
                   //PathData - command - valueFlags
                   //====================================================================================================================================
                   // also copy flagMode to pathDataPreBuf for use in specific case of waitFlag
                   FOR #tempFlagCtr := 1 TO "LKINCTRL_NO_OF_CMD_VALUEFLAGS" DO
                       #pathDataPreBuf.commands[#pathDataPreBuf.addPointer].valueFlags[#tempFlagCtr] := #statPathDataCommand.valueFlags[#tempFlagCtr];
                       // // change flagMode 3 to flagMode 2 as functionality is equal
                       // check for cmd to be flagOnly cmd
                       // check for cmd to implement flag and flagMode to be flagMode 3
                       IF #pathDataPreBuf.commands[#pathDataPreBuf.addPointer].cmdType = "LKINCTRL_CMD_FLAG_ONLY"
                           AND #pathDataPreBuf.commands[#pathDataPreBuf.addPointer].valueFlags[#tempFlagCtr].flag <> -1
                           AND #pathDataPreBuf.commands[#pathDataPreBuf.addPointer].valueFlags[#tempFlagCtr].flagMode = 3
                       THEN
                           // change flagMode 3 to flagMode 2
                           #pathDataPreBuf.commands[#pathDataPreBuf.addPointer].valueFlags[#tempFlagCtr].flagMode := 2;
                       END_IF;
                   END_FOR;

                   // skip lastPos calculation in case of wait time execution ==> old lastPos will be correct ==> use separation of config / motion cmd (flagOnly)
                   IF #statCmdIsMotionCmd THEN
                       //------------------------------------------------------------------------------------------
                       // Transform statLastPos into correct CS
                       //------------------------------------------------------------------------------------------
                       // TODO: Integrate InverseKinTrans into FC LKinCtrl_FrameTrans ?
                       IF #statPathDataCommand.cmdCoordinates.coordSystem = "CS_MCS"
                           AND #statCoordSystemOld <> "CS_MCS"
                       THEN
                           // Transform lastPos to MCS 
                           #instMC_InverseKinematicsTransformation(AxesGroup := #to_Kinematics,
                                                                   Enable := TRUE,
                                                                   Position := #statLastPos,
                                                                   CoordSystem := #statCoordSystemOld,
                                                                   LinkConstellation := #statLinkConstellation,
                                                                   ErrorId => #tempRetVal,
                                                                   AxesPosition => #statLastPos);

                       ELSIF #statPathDataCommand.cmdCoordinates.coordSystem <> "CS_MCS"
                           AND #statCoordSystemOld = "CS_MCS"
                       THEN
                           // Transform lastPos to target CS
                           #instMC_KinematicsTransformation(AxesGroup := #to_Kinematics,
                                                            Enable := TRUE,
                                                            AxesPosition := #statLastPos,
                                                            CoordSystem := #statPathDataCommand.cmdCoordinates.coordSystem,
                                                            ErrorId => #tempRetVal,
                                                            Position => #statLastPos,
                                                            LinkConstellation => #statLinkConstellation);

                       ELSE
                           // FR 26.03.2020: Updated FrameTrans 
                           // Transform LastPos to correct CS
                           "LKinCtrl_FrameTrans"(coordSystem := #statPathDataCommand.cmdCoordinates.coordSystem, // Actual/Target CS
                                                 coordSystemOld := #statCoordSystemOld, // Last CS
                                                 OCSFrames := #OCSFrames, // OCS frames
                                                 position := #statLastPos); // Position to be transformed
                       END_IF;

                       // Check if KinTrans FBs returned no error
                       IF #tempRetVal = 16#0 THEN
                           // Update old CS
                           #statCoordSystemOld := #statPathDataCommand.cmdCoordinates.coordSystem;

                           //------------------------------------------------------------------------------------------
                           // Update linkConstellation
                           //------------------------------------------------------------------------------------------
                           // LinkConstellation can only be set at sPTP command in WCS/OCS
                           IF #statPathDataCommand.cmdCoordinates.coordSystem <> "CS_MCS"
                               AND #statPathDataCommand.cmdParameters.moveDirectParameters.linkConstellation <> 16#FFFF_FFFF
                               AND (#statPathDataCommand.cmdType = "LKINCTRL_MC_MOVEDIRECTABS"
                               OR #statPathDataCommand.cmdType = "LKINCTRL_MC_MOVEDIRECTREL")
                           THEN
                               // LinkConstellation is changed
                               #statLinkConstellation := DWORD_TO_DINT(#statPathDataCommand.cmdParameters.moveDirectParameters.linkConstellation);
                           END_IF;

                           //------------------------------------------------------------------------------------------
                           // Update PositionMode
                           //------------------------------------------------------------------------------------------
                           // PositionMode is only valid for absolute SPTP command in WCS/OCS
                           IF #statPathDataCommand.cmdCoordinates.coordSystem <> "CS_MCS"
                               AND #statPathDataCommand.cmdParameters.moveDirectParameters.positionMode = 2 // Relative A coordinate
                               AND #statPathDataCommand.cmdType = "LKINCTRL_MC_MOVEDIRECTABS"
                           THEN
                               // Calc correct orientation position
                               #statLastPos[4] := #statLastPos[4] + #statPathDataCommand.cmdCoordinates.cartesianPosition.a;
                           END_IF;

                           //------------------------------------------------------------------------------------------
                           // ParameterValid bit check
                           //------------------------------------------------------------------------------------------
                           // added FR: 2020/04/03
                           "LKinCtrl_EvaluateParamValidBits"(parameterValidBits := #statParameterValid,
                                                             lastPos := #statLastPos,
                                                             errorMessage => #statDebugMessage,
                                                             command := #statPathDataCommand);

                           // Caclulation of resulting last position after command
                           //====================================================================================================================================
                           #statRetValLastPos := "LKinCtrl_CalcResultingPos"(cmdType := #statPathDataCommand.cmdType,
                                                                             cartesianPos := #statPathDataCommand.cmdCoordinates.cartesianPosition,
                                                                             circleParameters := #statPathDataCommand.cmdParameters.circleParameters,
                                                                             errorMessage => #statDebugMessage,
                                                                             lastPos := #statLastPos,
                                                                             lastAuxPoint := #statAuxPoint);

                           // check for error in last position calculation
                           IF #statRetValLastPos <> 16#0 THEN
                               // set error status
                               #statErrorAutoCleared := TRUE;
                               #statStatus := #ERR_LASTPOS_CALCULATION;
                           END_IF;

                       ELSE
                           // Error in KinTrans FBs
                           // set error status
                           #statErrorAutoCleared := TRUE;
                           #statStatus := #tempRetVal;
                       END_IF;

                   END_IF;

                   // PathData Blending at start of path
                   IF (#statPathDataPointers.retrievePointer = 1) AND
                       (#initPathTransition = 1)
                   THEN
                       #pathDataPreBuf.commands[#pathDataPreBuf.addPointer].cmdParameters.bufferMode := #initBufferMode;
                       #pathDataPreBuf.commands[#pathDataPreBuf.addPointer].cmdParameters.transitionParameters := #initTransitionParameter;
                   END_IF;

                   // increment PathDataPreBuf addPointer for next copy procedure
                   // also implement restart of pointer (1..constant)
                   IF #pathDataPreBuf.addPointer < "LKINCTRL_NO_OF_PATHDATA_PREBUFFER_ELEMENTS" THEN
                       #pathDataPreBuf.addPointer += 1;
                   ELSE
                       #pathDataPreBuf.addPointer := 1;
                       #pathDataPreBuf.addPointerRestarted := TRUE;
                   END_IF;
               END_REGION COPY_CMD_REGULAR

               // Go to copy cmd
               #statStateMachine := #GET_CMD;
           END_IF;


           // =======================================================================================================  
           // Contour offset is handled in the following regions / states
           // =======================================================================================================  
           REGION CONTOUR_OFFSET

               // STATE: CHECK_NEXT_CMD
               // =======================================================================================================  
               // CHECK_NEXT_CMD: Check next command for contour offset (#statPathCmdOffCompIn.nextCommand)
               // Next state: OFFSET_CALC / SEARCH_NBO
               IF #statStateMachine = #CHECK_NEXT_CMD THEN
                   REGION CHECK_NEXT_CMD
                       // Check if current command has length 0.0 --> Copy without contour offset
                       // else use as nextCmd & search NBO
                       // Transform lastPos to correct CS
                       "LKinCtrl_FrameTrans"(coordSystem := #statPathDataCommand.cmdCoordinates.coordSystem,
                                             coordSystemOld := #statCoordSystemOld,
                                             OCSFrames := #OCSFrames,
                                             position := #statLastPos);

                       // Update old CS
                       #statCoordSystemOld := #statPathDataCommand.cmdCoordinates.coordSystem;

                       // ParameterValid bit check
                       "LKinCtrl_EvaluateParamValidBits"(parameterValidBits := #statParameterValid,
                                                         lastPos := #statLastPos,
                                                         errorMessage => #statDebugMessage,
                                                         command := #statPathDataCommand);

                       // implement CM3 ==> CM1 conversion here
                       #statRetValCircModeConv := "LKinCtrl_ConvCircMode3To1"(coordinates := #statPathDataCommand.cmdCoordinates.cartesianPosition,
                                                                              errorMessage => #statDebugMessage,
                                                                              lastPos := #statLastPos,
                                                                              cmdType := #statPathDataCommand.cmdType,
                                                                              circleParameters := #statPathDataCommand.cmdParameters.circleParameters);

                       // Check if cmd has 0.0 length
                       "LKinCtrl_CheckForCmdLengthZero"(lastPos := #statLastPos,
                                                        commandLengthIsZero => #tempCmdLengthIsZero,
                                                        command := #statPathDataCommand);

                       // check for command length to be zero
                       IF #tempCmdLengthIsZero = FALSE THEN
                           // Comd is not length 0.0

                           // Calc resulting pos to use for searching NBO
                           #statRetValLastPos := "LKinCtrl_CalcResultingPos"(cmdType := #statPathDataCommand.cmdType,
                                                                             cartesianPos := #statPathDataCommand.cmdCoordinates.cartesianPosition,
                                                                             circleParameters := #statPathDataCommand.cmdParameters.circleParameters,
                                                                             errorMessage => #statDebugMessage,
                                                                             lastAuxPoint := #statAuxPoint,
                                                                             lastPos := #statLastPos);


                           // Use as next cmd
                           // set first condition bit to abort loop
                           #tempValidNextCmdFound := TRUE;
                           #statDebugNextCmdFound := #statPathDataPointers.retrievePointer;

                           // check for command to be END_OFFSET_COMP command
                           IF #statPathDataCommand.cmdType = "LKINCTRL_CONFIG_END_OFFSET_COMP"
                               OR #statPathDataCommand.cmdType = -1
                           THEN
                               // transfer no command for end of compensation
                               #statPathCmdOffCompIn.nextCommand.cmdType := -1;
                               // transfer no command for end of compensation
                               #statPathCmdOffCompIn.nextButOneCommand.cmdType := -1;
                               #tempValidNextButOneCmdFound := TRUE;
                               // Go to next state --> No need to search NBO
                               #statStateMachine := #OFFSET_CALC;
                           ELSE
                               // copy 'next' cmd to next(ButOne)Command input
                               #statPathCmdOffCompIn.nextCommand := #statPathDataCommand;
                               // Go to next state
                               #statStateMachine := #SEARCH_NBO;
                           END_IF;

                       ELSE
                           // command has no length --> RelCmd with 0.0 or AbsCmd with same target
                           // copy command as usual without calling any contour offset calculation functions
                           REGION COPY_LENGTH_0_CMD
                               //PathData - command - cmdType
                               #pathDataPreBuf.commands[#pathDataPreBuf.addPointer].cmdType := #statPathDataCommand.cmdType;

                               //PathData - command - cmdID
                               #pathDataPreBuf.commands[#pathDataPreBuf.addPointer].cmdID := #statPathDataPointers.retrievePointer + #statNoRestarts * INT_TO_DINT("LKINCTRL_NO_OF_PATHDATA_ELEMENTS_ADVANCED");

                               //PathData - command - cmdName
                               #pathDataPreBuf.commands[#pathDataPreBuf.addPointer].cmdName := #statPathDataCommand.cmdName;

                               //PathData - command - cmdCoordinates
                               //====================================================================================================================================
                               //PathData - command - cmdCoordinates - absolutePosition[1..4]
                               IF #statOffsetCompFirstCmd = FALSE AND #statPathDataCommand.cmdType = "LKINCTRL_MC_MOVELINEARABS" THEN
                                   // Use compensated coordinates for multiple zero length commands in a row
                                   #pathDataPreBuf.commands[#pathDataPreBuf.addPointer].cmdCoordinates.absolutePosition[1] := #statPathCmdOffCompIn.currentPos.positionAbsoluteRadComp.x;
                                   #pathDataPreBuf.commands[#pathDataPreBuf.addPointer].cmdCoordinates.absolutePosition[2] := #statPathCmdOffCompIn.currentPos.positionAbsoluteRadComp.y;
                                   #pathDataPreBuf.commands[#pathDataPreBuf.addPointer].cmdCoordinates.absolutePosition[3] := #statPathCmdOffCompIn.currentPos.positionAbsoluteRadComp.z;
                                   #pathDataPreBuf.commands[#pathDataPreBuf.addPointer].cmdCoordinates.absolutePosition[4] := #statPathCmdOffCompIn.currentPos.positionAbsoluteRadComp.a;
                               ELSE
                                   #pathDataPreBuf.commands[#pathDataPreBuf.addPointer].cmdCoordinates.absolutePosition[1] := #statPathDataCommand.cmdCoordinates.cartesianPosition.x;
                                   #pathDataPreBuf.commands[#pathDataPreBuf.addPointer].cmdCoordinates.absolutePosition[2] := #statPathDataCommand.cmdCoordinates.cartesianPosition.y;
                                   #pathDataPreBuf.commands[#pathDataPreBuf.addPointer].cmdCoordinates.absolutePosition[3] := #statPathDataCommand.cmdCoordinates.cartesianPosition.z;
                                   #pathDataPreBuf.commands[#pathDataPreBuf.addPointer].cmdCoordinates.absolutePosition[4] := #statPathDataCommand.cmdCoordinates.cartesianPosition.a;
                               END_IF;

                               //PathData - command - cmdCoordinates - coordSystem
                               #pathDataPreBuf.commands[#pathDataPreBuf.addPointer].cmdCoordinates.coordSystem := #statPathDataCommand.cmdCoordinates.coordSystem;

                               //PathData - command - cmdParameters
                               //====================================================================================================================================
                               //PathData - command - cmdParameters - pathDynamics
                               #pathDataPreBuf.commands[#pathDataPreBuf.addPointer].cmdParameters.pathDynamics := #statPathDataCommand.cmdParameters.pathDynamics;

                               //PathData - command - cmdParameters - orientationDirection
                               #pathDataPreBuf.commands[#pathDataPreBuf.addPointer].cmdParameters.orientationDirection := #statPathDataCommand.cmdParameters.orientationDirection;

                               //PathData - command - cmdParameters - bufferMode
                               #pathDataPreBuf.commands[#pathDataPreBuf.addPointer].cmdParameters.bufferMode := #statPathDataCommand.cmdParameters.bufferMode;

                               //PathData - command - cmdParameters - transitionParameters
                               #pathDataPreBuf.commands[#pathDataPreBuf.addPointer].cmdParameters.transitionParameters[1] := #statPathDataCommand.cmdParameters.transitionParameters[1];

                               //PathData - command - cmdParameters - dynamicAdaption
                               #pathDataPreBuf.commands[#pathDataPreBuf.addPointer].cmdParameters.dynamicAdaption := #statPathDataCommand.cmdParameters.dynamicAdaption;

                               //PathData - command - setFlags
                               //====================================================================================================================================
                               // also copy flagMode to pathDataPreBuf for use in specific case of waitFlag
                               FOR #tempFlagCtr := 1 TO "LKINCTRL_NO_OF_CMD_SETFLAGS" DO
                                   #pathDataPreBuf.commands[#pathDataPreBuf.addPointer].setFlags[#tempFlagCtr] := #statPathDataCommand.setFlags[#tempFlagCtr];
                                   // // change flagMode 3 to flagMode 2 as functionality is equal
                                   // check for cmd to be flagOnly cmd
                                   // check for cmd to implement flag and flagMode to be flagMode 3
                                   IF #pathDataPreBuf.commands[#pathDataPreBuf.addPointer].cmdType = "LKINCTRL_CMD_FLAG_ONLY"
                                       AND #pathDataPreBuf.commands[#pathDataPreBuf.addPointer].setFlags[#tempFlagCtr].flag <> -1
                                       AND #pathDataPreBuf.commands[#pathDataPreBuf.addPointer].setFlags[#tempFlagCtr].flagMode = 3
                                   THEN
                                       // change flagMode to flagMode 1
                                       #pathDataPreBuf.commands[#pathDataPreBuf.addPointer].setFlags[#tempFlagCtr].flagMode := 2;
                                   END_IF;
                               END_FOR;

                               //PathData - command - valueFlags
                               //====================================================================================================================================
                               // also copy flagMode to pathDataPreBuf for use in specific case of waitFlag
                               FOR #tempFlagCtr := 1 TO "LKINCTRL_NO_OF_CMD_VALUEFLAGS" DO
                                   #pathDataPreBuf.commands[#pathDataPreBuf.addPointer].valueFlags[#tempFlagCtr] := #statPathDataCommand.valueFlags[#tempFlagCtr];
                                   // // change flagMode 3 to flagMode 2 as functionality is equal
                                   // check for cmd to be flagOnly cmd
                                   // check for cmd to implement flag and flagMode to be flagMode 3
                                   IF #pathDataPreBuf.commands[#pathDataPreBuf.addPointer].cmdType = "LKINCTRL_CMD_FLAG_ONLY"
                                       AND #pathDataPreBuf.commands[#pathDataPreBuf.addPointer].valueFlags[#tempFlagCtr].flag <> -1
                                       AND #pathDataPreBuf.commands[#pathDataPreBuf.addPointer].valueFlags[#tempFlagCtr].flagMode = 3
                                   THEN
                                       // change flagMode to flagMode 1
                                       #pathDataPreBuf.commands[#pathDataPreBuf.addPointer].valueFlags[#tempFlagCtr].flagMode := 2;
                                   END_IF;

                               END_FOR;

                               // increase addPointer after copy of command for next command
                               IF #pathDataPreBuf.addPointer < "LKINCTRL_NO_OF_PATHDATA_PREBUFFER_ELEMENTS" THEN
                                   #pathDataPreBuf.addPointer += 1;
                               ELSE
                                   #pathDataPreBuf.addPointer := 1;
                                   #pathDataPreBuf.addPointerRestarted := TRUE;
                               END_IF;

                           END_REGION COPY_REL_0_CMD

                           // Go to next state
                           #statStateMachine := #OFFSET_CALC;

                       END_IF;
                   END_REGION CHECK_NEXT_CMD
               END_IF;


               // STATE: SEARCH_NBO
               // =======================================================================================================  
               // SEARCH_NBO: Search forward in path data for contour offset next but one command (#statPathCmdOffCompIn.nextButOneCommand)
               // Next state: OFFSET_CALC
               IF #statStateMachine = #SEARCH_NBO THEN
                   REGION SEARCH_NBO
                       // find valid nextCmd and nextButOneCmd (input) data
                       // ---------------------------------------------------
                       // Init last pos and old coord system
                       #statNBOLastPos := #statLastPos;
                       #tempNBOCoordSystemOld := #statCoordSystemOld;

                       IF #statSearchNBOAborted = FALSE THEN
                           // initially set pointer increase counter to 1
                           #statRetrievePointerIncCtr := 1;
                       ELSE
                           // Reset abort bit but keep RetreivePointerIncCounter the same
                           #statSearchNBOAborted := FALSE;
                       END_IF;

                       // Use repeat to search in path data for next valid command
                       REPEAT

                           // Check pointers also for not ringBuffer or ignore add pointer
                           // Added FR 22.05.2019
                           IF #statPathDataPointers.ignoreAddPointer THEN
                               // No ring buffer
                               // Check index to be lower than max path data length 
                               IF #statPathDataType = "LKINCTRL_PATHDATA_TYPE_REDUCED" THEN
                                   #tempIndexOk := #statPathDataPointers.retrievePointer + #statRetrievePointerIncCtr <= "LKINCTRL_NO_OF_PATHDATA_ELEMENTS_REDUCED";
                               ELSIF #statPathDataType = "LKINCTRL_PATHDATA_TYPE_NORMAL" THEN
                                   #tempIndexOk := #statPathDataPointers.retrievePointer + #statRetrievePointerIncCtr <= "LKINCTRL_NO_OF_PATHDATA_ELEMENTS";
                               ELSIF #statPathDataType = "LKINCTRL_PATHDATA_TYPE_ADVANCED" THEN
                                   #tempIndexOk := #statPathDataPointers.retrievePointer + #statRetrievePointerIncCtr <= "LKINCTRL_NO_OF_PATHDATA_ELEMENTS_ADVANCED";
                               END_IF;
                           ELSE
                               // Ring buffer
                               // Added JR 13.05.2019 
                               // If index overflows then calc offset to point to first index
                               IF #statPathDataPointers.retrievePointer + #statRetrievePointerIncCtr > "LKINCTRL_NO_OF_PATHDATA_ELEMENTS_ADVANCED" THEN
                                   // Set statRetrievePointerIncCtr
                                   #statRetrievePointerIncCtr := 1 - #statPathDataPointers.retrievePointer;
                               END_IF;

                               // Condition if (#statPathDataPointers.retrievePointer + #statRetrievePointerIncCtr) > 1
                               #tempIndexOk :=
                               ((#statPathDataPointers.retrievePointer + #statRetrievePointerIncCtr) <= #statPathDataPointers.addPointer)
                               OR (((#statPathDataPointers.retrievePointer + #statRetrievePointerIncCtr) > #statPathDataPointers.addPointer)
                               AND #statPathDataPointers.addPointerRestarted);
                           END_IF;

                           // Copy path data command
                           // 2019.03.28 FR: Get last command
                           IF (#statPathDataPointers.retrievePointer + #statRetrievePointerIncCtr) >= 1
                               AND #tempIndexOk
                           THEN
                               // Get path data command and previous path data command
                               #tempRetVal := "LKinCtrl_GetPathDataCmd"(pathDataType := #statPathDataType,
                                                                        index := #statPathDataPointers.retrievePointer + #statRetrievePointerIncCtr,
                                                                        pathDataReduced := #tempPathData_reduced,
                                                                        pathData := #tempPathData,
                                                                        pathDataAdvanced := #tempPathData_advanced,
                                                                        pathDataCommand => #statPathCmdNBOCheck,
                                                                        parameterValid => #tempParameterValidNBO);


                               // Check if index is not ok and not ring buffer
                               // --> End of path data is reached and Next or NBO was not found 
                               // --> Set the corresponding cmd to -1 to end offset correctly 
                           ELSIF #tempIndexOk = FALSE
                               AND #statPathDataPointers.ignoreAddPointer
                           THEN
                               IF #tempValidNextCmdFound THEN
                                   // set NBO to -1
                                   // transfer no command for end of compensation
                                   #statPathCmdOffCompIn.nextButOneCommand.cmdType := -1;
                                   #tempValidNextButOneCmdFound := TRUE;
                               ELSE
                                   // set Next and NBO to -1
                                   // transfer no command for end of compensation
                                   #statPathCmdOffCompIn.nextCommand.cmdType := -1;
                                   #tempValidNextCmdFound := TRUE;
                                   // transfer no command for end of compensation
                                   #statPathCmdOffCompIn.nextButOneCommand.cmdType := -1;
                                   #tempValidNextButOneCmdFound := TRUE;
                               END_IF;
                               // Exit repeat
                               EXIT;

                               // Index is not valid and ringbuffer active --> Check for new command 
                           ELSE
                               // Exit repeat loop and check again in next cycle
                               // memorize abort
                               #statSearchNBOAborted := TRUE;
                               EXIT;
                           END_IF;

                           // preCheck sequence for comamnd to have length of zero
                           #tempCmdLengthIsZero := FALSE;

                           // Command was copied --> Check if valid for NBO
                           IF #statPathCmdNBOCheck.cmdActivated THEN
                               // Valid
                               // Check for length 0.0
                               // Transform lastPos to correct CS
                               "LKinCtrl_FrameTrans"(coordSystem := #statPathCmdNBOCheck.cmdCoordinates.coordSystem,
                                                     coordSystemOld := #tempNBOCoordSystemOld,
                                                     OCSFrames := #OCSFrames,
                                                     position := #statNBOLastPos);

                               // Update old CS
                               #tempNBOCoordSystemOld := #statPathCmdNBOCheck.cmdCoordinates.coordSystem;

                               // ParameterValid bit check
                               "LKinCtrl_EvaluateParamValidBits"(parameterValidBits := #tempParameterValidNBO,
                                                                 lastPos := #statNBOLastPos,
                                                                 errorMessage => #statDebugMessage,
                                                                 command := #statPathCmdNBOCheck);

                               // implement CM3 ==> CM1 conversion here
                               #statRetValCircModeConv := "LKinCtrl_ConvCircMode3To1"(coordinates := #statPathCmdNBOCheck.cmdCoordinates.cartesianPosition,
                                                                                      errorMessage => #statDebugMessage,
                                                                                      lastPos := #statNBOLastPos,
                                                                                      cmdType := #statPathCmdNBOCheck.cmdType,
                                                                                      circleParameters := #statPathCmdNBOCheck.cmdParameters.circleParameters);

                               // Check if cmd has 0.0 length
                               "LKinCtrl_CheckForCmdLengthZero"(lastPos := #statNBOLastPos,
                                                                commandLengthIsZero => #tempCmdLengthIsZero,
                                                                command := #statPathCmdNBOCheck);

                               IF #tempCmdLengthIsZero = FALSE THEN
                                   // Has length
                                   // Check if valid
                                   // set condition bit to abort loop
                                   #tempValidNextButOneCmdFound := TRUE;
                                   #statDebugNextButOneCmdFound := #statPathDataPointers.retrievePointer + #statRetrievePointerIncCtr;

                                   // check for command to be END_OFFSET_COMP command
                                   IF #statPathCmdNBOCheck.cmdType = "LKINCTRL_CONFIG_END_OFFSET_COMP"
                                       OR #statPathCmdNBOCheck.cmdType = -1
                                   THEN
                                       // transfer no command for end of compensation
                                       #statPathCmdOffCompIn.nextButOneCommand.cmdType := -1;
                                   ELSE
                                       // copy 'next' cmd to nextButOneCommand input
                                       #statPathCmdOffCompIn.nextButOneCommand := #statPathCmdNBOCheck;
                                   END_IF;
                               ELSE
                                   // Is 0.0 length cmd --> Not valid for NBO --> Search continues
                                   // increase set pointer increase counter to check next element
                                   #statRetrievePointerIncCtr += 1;
                               END_IF;

                           ELSE
                               // Cmd deactivated --> Not valid
                               // increase set pointer increase counter to check next element
                               #statRetrievePointerIncCtr += 1;
                           END_IF;

                       UNTIL #tempValidNextButOneCmdFound END_REPEAT;

                       // If both cmds were found and no abort then go to offset calc
                       IF #tempValidNextButOneCmdFound AND NOT #statSearchNBOAborted THEN
                           // Go to OffsetCalc
                           #statStateMachine := #OFFSET_CALC;

                           // reset variable for first offset command
                           #statOffsetCompFirstCmd := FALSE;
                       END_IF;
                   END_REGION SEARCH_NBO
               END_IF;

               // STATE: OFFSET_CMD
               // =======================================================================================================   
               // OFFSET_CMD: Copy offset command
               IF #statStateMachine = #OFFSET_CALC THEN
                   REGION OFFSET_CALC
                       // Offset Compensation Calculation
                       //====================================================================================================================================
                       // prepare data for offset calculation ==> only use original commands (source Pathdata !)

                       // check for command length not to be zero
                       IF #tempCmdLengthIsZero = FALSE THEN

                           // run offset caclulation
                           #statRetValOffsetComp := "LKinCtrl_OffsetContour"(toolLength := #statToolLength,
                                                                             toolRadius := #statToolRadius,
                                                                             pathPlane := #statPathPlane,
                                                                             compensationDirection := #statCompDirection,
                                                                             pathDataIn := #statPathCmdOffCompIn,
                                                                             pathDataOut := #statPathCmdOffCompOut);

                           // check for errors in offset compensation calculation
                           IF #statRetValOffsetComp.returnValue <> 16#0 THEN
                               #statErrorAutoCleared := TRUE;
                               #statStatus := #statRetValOffsetComp.returnValue;
                           ELSE
                               // use nextPositionAbsolute from last calc as currentPositionAbsolute for next calc
                               #statPathCmdOffCompIn.currentPos.positionAbsolute := #statPathCmdOffCompOut.nextPositionAbsolute;
                               #statPathCmdOffCompIn.currentPos.positionAbsoluteRadComp := #statPathCmdOffCompOut.nextPositionAbsoluteRadComp;

                               // use results of offset compensation calculation
                               // check for compensated nextCmd to be available
                               IF #statPathCmdOffCompOut.nextCommand.cmdType <> -1 THEN
                                   //PathData - command - cmdID
                                   #pathDataPreBuf.commands[#pathDataPreBuf.addPointer].cmdID := #statPathDataPointers.retrievePointer + #statNoRestarts * INT_TO_DINT("LKINCTRL_NO_OF_PATHDATA_ELEMENTS_ADVANCED");

                                   // copy next cmd data (OUT) - compensated (new calculated data)
                                   "LKinCtrl_ConvElements_PathDataToPathData_PreBuf"(copyCompensatedParametes := TRUE,
                                                                                     copyTransitionParameters := FALSE, //true ,
                                                                                     copyFlags := TRUE,
                                                                                     pathDataElement := #statPathCmdOffCompOut.nextCommand,
                                                                                     pathDataPreBufElement := #pathDataPreBuf.commands[#pathDataPreBuf.addPointer],
                                                                                     pathDataName := #statPathDataName);

                                   // Added FR 22.05.2019: Set ParameterValid bits true
                                   FOR #tempCtr := 1 TO "LKINCTRL_NO_OF_VALID_BITS" DO
                                       #pathDataPreBuf.commands[#pathDataPreBuf.addPointer].parameterValid[#tempCtr] := TRUE;
                                   END_FOR;

                                   // increase addPointer after copy of command for next command
                                   IF #pathDataPreBuf.addPointer < "LKINCTRL_NO_OF_PATHDATA_PREBUFFER_ELEMENTS" THEN
                                       #pathDataPreBuf.addPointer += 1;
                                   ELSE
                                       #pathDataPreBuf.addPointer := 1;
                                       #pathDataPreBuf.addPointerRestarted := TRUE;
                                   END_IF;

                                   // write transitionParameters of nextButOneCmd result to next but one command
                                   #pathDataPreBuf.commands[#pathDataPreBuf.addPointer].cmdParameters.transitionParameters := #statPathCmdOffCompOut.nextButOneCommand.transitionParameter;
                               ELSE
                                   ; // Invalid command -> nothing to copy
                               END_IF;

                               // check if there is an additional intermediate command
                               IF (#statPathCmdOffCompOut.intermediateCommand.cmdType > 0) THEN

                                   // copy intermediate cmd to PathData_PreBuf - no flags
                                   "LKinCtrl_ConvElements_PathDataToPathData_PreBuf"(copyCompensatedParametes := TRUE,
                                                                                     copyTransitionParameters := FALSE,
                                                                                     copyFlags := FALSE,
                                                                                     pathDataElement := #statPathCmdOffCompOut.intermediateCommand,
                                                                                     pathDataPreBufElement := #pathDataPreBuf.commands[#pathDataPreBuf.addPointer],
                                                                                     pathDataName := #statPathDataName);

                                   //PathData - command - cmdID
                                   // set intermediate commands cmdID to cmdID of following command ==> flag handling similar to transitionParameter
                                   #pathDataPreBuf.commands[#pathDataPreBuf.addPointer].cmdID := (#statPathDataPointers.retrievePointer + 1) + #statNoRestarts * INT_TO_DINT("LKINCTRL_NO_OF_PATHDATA_ELEMENTS_ADVANCED");

                                   // added FR: 11.07.2019: Set ParameterValid bits true
                                   FOR #tempCtr := 1 TO "LKINCTRL_NO_OF_VALID_BITS" DO
                                       #pathDataPreBuf.commands[#pathDataPreBuf.addPointer].parameterValid[#tempCtr] := TRUE;
                                   END_FOR;

                                   // mark intermediate commands to except them from flag for remaining distance
                                   #pathDataPreBuf.commands[#pathDataPreBuf.addPointer].isIntermediateCmd := TRUE;

                                   // increase addPointer after copy of command for next command
                                   IF #pathDataPreBuf.addPointer < "LKINCTRL_NO_OF_PATHDATA_PREBUFFER_ELEMENTS" THEN
                                       #pathDataPreBuf.addPointer += 1;
                                   ELSE
                                       #pathDataPreBuf.addPointer := 1;
                                       #pathDataPreBuf.addPointerRestarted := TRUE;
                                   END_IF;

                               ELSE
                                   ; // No intermediate cmd -> do nothing
                               END_IF;
                           END_IF;

                       ELSE
                           ; // do nothing --> Command was already copied
                       END_IF;

                   END_REGION OFFSET_CALC

                   // Go to copy cmd
                   #statStateMachine := #GET_CMD;
               END_IF;
           END_REGION CONTOUR_OFFSET

       END_REGION PATHDATA_PREBUFFERING


       REGION PATHDATA_PREBUFFERED_COMPLETELY
           // STATE: PATHDATA_PREBUFFERED_COMPLETELY
           // =======================================================================================================      
           // PATHDATA_PREBUFFERED_COMPLETELY: Disabling, e.g. closing connections, etc.
           IF #statStateMachine = #PATHDATA_PREBUFFERED_COMPLETELY
               // AND #statDebugState = TRUE
           THEN

               // reset  variable for single step debugging of states
               #statDebugState := FALSE;

               // Added FR 2019.03.28 // Reworked 08.04.2020
               // REGION GET_LAST_CMD_TYPE
               //
               // Always get last cmd id from preBuffered
               // --> Deactivated commands do not appear in preBuffered anyway
               // --> No need to check config cmds as they also do not appear --> Output LastCmdIsConfigCmd is not even needed / used in MovePath
               // --> Last cmdType equals cmdID element
               // --> LastCmdId is checked in MovePath if all commands are executed by Executer 
               // --> Condition: LastCmdIdPathdata = PathDataElementPreBuffered.cmdId --> Check if all commands we added are executed
               // --> Problems: how to check if empty pathdata is connected?
               //               How to check if pathData with only deactivated cmds (and one -1) is connected 
               //               Or only config commands, ...
               //   ==> in all cases not a single command was added to preBuffer
               //   
               // Use bit to check if at least one command was added 
               IF #statCmdAdded THEN
                   // At least one command was added to PreBuffered PathData
                   // --> Use CmdId from PreBuffer to get statLastCmdId
                   // Prebuffered cmd at last addPointer index has last cmdID
                   IF (#pathDataPreBuf.addPointer - 1) > 0 THEN
                       #statLastCmdIdPathdata := #pathDataPreBuf.commands[#pathDataPreBuf.addPointer - 1].cmdID;
                   ELSE
                       #statLastCmdIdPathdata := #pathDataPreBuf.commands["LKINCTRL_NO_OF_PATHDATA_PREBUFFER_ELEMENTS"].cmdID;
                   END_IF;
               ELSE
                   // No command was added to PreBuffered PathData
                   // --> statLastCmdId = 0 
                   #statLastCmdIdPathdata := 0;
               END_IF;
           END_IF;
       END_REGION PATHDATA_PREBUFFERED_COMPLETELY


       REGION DISABLE_STATE
           // STATE: DISABLE_STATE
           // =======================================================================================================      
           // DISABLE_STATE: Disabling, e.g. closing connections, etc.
           IF #statStateMachine = #DISABLE_STATE
               // AND #statDebugState = TRUE
           THEN
               // reset  variable for single step debugging of states
               #statDebugState := FALSE;

               // reset variables before disabling -> will be reset at next enable
               IF TypeOf(#pathData) = LKinCtrl_typePathData_advanced THEN
                   #tempPathData_advanced ?= #pathData;

                   // added 2020.02.07 DF/FR: Reset retrieve pointer in PathData
                   #tempPathData_advanced<?OpDeref?>.pointers.retrievePointer := 0;
                   #statPathDataPointers := #tempPathData_advanced<?OpDeref?>.pointers;
               END_IF;

               // set statDisablingCompleted for deactivation of FB below
               #statDisablingCompleted := TRUE;

           END_IF;
       END_REGION DISABLE_STATE


   END_REGION STATE_MACHINE

   // reset of #pathDataPreBuf.addPointerRestarted in MovePath (called in every cycle)

   REGION OUTPUTS
       // Write outputs
       IF (#statDisablingCompleted = TRUE) THEN
           // Reset outputs if disabling completed
           #statValid := FALSE;
           #statBusy := FALSE;
           #statError := FALSE;
           #statErrorUserCleared := FALSE;
           // #statErrorAutoCleared := FALSE;
           #statStatus := #STATUS_NO_CALL;
           // TODO: Reset application specific outputs

       ELSIF (#statErrorUserCleared = TRUE) AND (#statError = FALSE) THEN
           // Error can only be cleared by user; rising edge at enable input is needed to continue 
           #statValid := FALSE;
           #statBusy := FALSE;
           #statError := TRUE;
           #statStateMachine := #NO_PROCESSING; // Switch state machine to "no processing"

       ELSIF (#statErrorAutoCleared = TRUE) AND (#statError = FALSE) THEN
           // Error can be reset by FB automatically  
           #statValid := FALSE;
           #statBusy := TRUE;
           #statError := TRUE;
           #statStateMachine := #NO_PROCESSING; // Switch state machine to "no processing"

       ELSIF (#statErrorAutoCleared = FALSE) AND (#statErrorUserCleared = FALSE) AND (#statError = TRUE) THEN
           // If autocleared error is acknowledged
           #statValid := TRUE;
           #statBusy := TRUE;
           #statError := FALSE;
           #statStatus := #STATUS_SUBSEQUENT_CALL;
       END_IF;

       // Copy pointers back to connected path data 
       IF #statPathDataType = "LKINCTRL_PATHDATA_TYPE_ADVANCED" THEN
           #tempPathData_advanced<?OpDeref?>.pointers := #statPathDataPointers;
       ELSE
           ; // No pointers outside --> Do nothing
       END_IF;

       // Write static values to outputs
       #valid := #statValid;
       #busy := #statBusy;
       #error := #statError;
       #status := #statStatus;
       // Write application specific static values to outputs
       #lastCmdIdPathData := #statLastCmdIdPathdata;
       #pathDataRetrievePointer := #statPathDataPointers.retrievePointer;
       #preprocessingStop := #statPathDataPointers.preprocessingStop;
   END_REGION OUTPUTS

   // =================================================================================================================
   // End of Function Block: LKinCtrl_PreBuffer
   // =================================================================================================================
END_FUNCTION_BLOCK

